(* Logix 5000 project; controller NWGG 1756-L72 rev 35.12; software revision 35.00; part 14 of 19 *)
(* tags used below, declared in another part *)
   ALM_Air_Gate_Failed_Open_Bin0 : ALARM_DIGITAL;
   ALM_Air_Gate_Failed_Open_Bin1 : ALARM_DIGITAL;
   ALM_Air_Gate_Failed_Open_Bin10 : ALARM_DIGITAL;
   ALM_Air_Gate_Failed_Open_Bin11 : ALARM_DIGITAL;
   ALM_Air_Gate_Failed_Open_Bin12 : ALARM_DIGITAL;
   ALM_Air_Gate_Failed_Open_Bin13 : ALARM_DIGITAL;
   ALM_Air_Gate_Failed_Open_Bin14 : ALARM_DIGITAL;
   ALM_Air_Gate_Failed_Open_Bin15 : ALARM_DIGITAL;
   ALM_Air_Gate_Failed_Open_Bin16 : ALARM_DIGITAL;
   ALM_Air_Gate_Failed_Open_Bin2 : ALARM_DIGITAL;
   ALM_Air_Gate_Failed_Open_Bin5 : ALARM_DIGITAL;
   ALM_Air_Gate_Failed_Open_Bin6 : ALARM_DIGITAL;
   ALM_Air_Gate_Failed_Open_Bin7 : ALARM_DIGITAL;
   ALM_Air_Gate_Failed_Open_Bin8 : ALARM_DIGITAL;
   ALM_Air_Gate_Failed_Open_Bin9 : ALARM_DIGITAL;
   ALM_OVRAMP_Belt10 : ALARM_DIGITAL;
   ALM_OVRAMP_Belt11 : ALARM_DIGITAL;
   ALM_OVRAMP_Belt2 : ALARM_DIGITAL;
   ALM_OVRAMP_Belt3 : ALARM_DIGITAL;
   ALM_OVRAMP_Belt5 : ALARM_DIGITAL;
   ALM_OVRAMP_Belt6 : ALARM_DIGITAL;
   ALM_OVRAMP_Belt7 : ALARM_DIGITAL;
   ALM_OVRAMP_Belt8 : ALARM_DIGITAL;
   ALM_OVRAMP_Belt9 : ALARM_DIGITAL;
   ALM_PLUG_Belt1 : ALARM_DIGITAL;
   ALM_PLUG_Belt10 : ALARM_DIGITAL;
   ALM_PLUG_Belt11 : ALARM_DIGITAL;
   ALM_PLUG_Belt2 : ALARM_DIGITAL;
   ALM_PLUG_Belt3 : ALARM_DIGITAL;
   ALM_PLUG_Belt5 : ALARM_DIGITAL;
   ALM_PLUG_Belt6 : ALARM_DIGITAL;
   ALM_PLUG_Belt7 : ALARM_DIGITAL;
   ALM_PLUG_Belt8 : ALARM_DIGITAL;
   ALM_PLUG_Belt9 : ALARM_DIGITAL;
   ALM_SLP10_Belt1 : ALARM_DIGITAL;
   ALM_SLP10_Belt10 : ALARM_DIGITAL;
   ALM_SLP10_Belt11 : ALARM_DIGITAL;
   ALM_SLP10_Belt2 : ALARM_DIGITAL;
   ALM_SLP10_Belt3 : ALARM_DIGITAL;
   ALM_SLP10_Belt5 : ALARM_DIGITAL;
   ALM_SLP10_Belt6 : ALARM_DIGITAL;
   ALM_SLP10_Belt7 : ALARM_DIGITAL;
   ALM_SLP10_Belt8 : ALARM_DIGITAL;
   ALM_SLP10_Belt9 : ALARM_DIGITAL;
   ALM_SLP20_Belt1 : ALARM_DIGITAL;
   ALM_SLP20_Belt10 : ALARM_DIGITAL;
   ALM_SLP20_Belt11 : ALARM_DIGITAL;
   ALM_SLP20_Belt2 : ALARM_DIGITAL;
   ALM_SLP20_Belt3 : ALARM_DIGITAL;
   ALM_SLP20_Belt5 : ALARM_DIGITAL;
   ALM_SLP20_Belt6 : ALARM_DIGITAL;
   ALM_SLP20_Belt7 : ALARM_DIGITAL;
   ALM_SLP20_Belt8 : ALARM_DIGITAL;
   ALM_SLP20_Belt9 : ALARM_DIGITAL;
   ALM_WONT_START_Belt1 : ALARM_DIGITAL;
   ALM_WONT_START_Belt10 : ALARM_DIGITAL;
   ALM_WONT_START_Belt11 : ALARM_DIGITAL;
   ALM_WONT_START_Belt2 : ALARM_DIGITAL;
   ALM_WONT_START_Belt3 : ALARM_DIGITAL;
   ALM_WONT_START_Belt5 : ALARM_DIGITAL;
   ALM_WONT_START_Belt6 : ALARM_DIGITAL;
   ALM_WONT_START_Belt7 : ALARM_DIGITAL;
   ALM_WONT_START_Belt8 : ALARM_DIGITAL;
   ALM_WONT_START_Belt9 : ALARM_DIGITAL;
   Always_Off : BOOL;
   Andco_Rate : DINT;
   b3 : ALARM_DIGITAL;
   Batch_Status : DINT;
   BC_9_Interlock : BOOL;
   Belt : udt_Motor[16];
   Bin_Clean_Pause : BOOL;
   Bin_Loadout_Control : Loadout_Bin_Control[29];
   Bin_Transfer_Pause : BOOL;
   Bin_Treat_Pause : BOOL;
   Clean_Batch_Status : DINT;
   Concrete_Leg : udt_Motor;
   Config_Bin_Name : STRING;
   Config_Cancel_Bin : BOOL;
   Config_Class : STRING;
   Config_Clean_Delay_Start : REAL;
   Config_Clean_Delay_Stop : REAL;
   Config_Item_Number : STRING;
   Config_Name : STRING;
   Config_Pounds_Per_Inch : REAL;
   Config_Save_Bin : BOOL;
   Config_Treat_Delay_Start : REAL;
   Config_Treat_Delay_Stop : REAL;
   ConfigureIndex : DINT;
   Empty_String : STRING;
   IDX : DINT;
   Interlock_Not_Used : BOOL;
   loa : ALARM_DIGITAL;
   Loadout_Bin : udt_Loadout_Bin[29];
   Loadout_K_Valve : udt_Loadout_K_Valve[2];
   Man_Start_Stop_Allowed : BOOL;
   Manual_Mode : BOOL;
   Move_Bin_Config : BOOL;
   NA : BOOL;
   TMR_Max_Clean_Delay : TIMER;
   TMR_Max_Treat_Delay : TIMER;
   Transfer_Batch_Status : DINT;
   Treat_Batch_Status : DINT;
   Treater_Loadout : udt_Treater_Loadout;
   _700_AIR_GA : ALIAS FOR I8.3;
   _700G_CLOSE : ALIAS FOR O12.9;
   _700G_OPEN : ALIAS FOR O12.8;
   _701_AIR_GA : ALIAS FOR I8.5;
   Always_On : BOOL;
   Bin_Config : BOOL;
   CP_Remote_Air_Gate_On : DINT;
   CP_Remote_Air_Gate_Open_In : DINT;
   CP_Remote_Andoc_Out : udt_Andco_Remote_Out[32];
   CP_Remote_Belt_In : udt_Motor_Remote_In[10];
   CP_Remote_Belt_Start : DINT;
   I1_000_Bit00 : ALIAS FOR I1.0;
   I4_000_Bit11 : ALIAS FOR I4.11;
   I8_000_Bit08 : ALIAS FOR I8.8;
   I8_000_Bit09 : ALIAS FOR I8.9;
   I8_000_Bit10 : ALIAS FOR I8.10;
   I8_000_Bit11 : ALIAS FOR I8.11;
   O12_000_Bit10 : ALIAS FOR O12.10;
   O12_000_Bit11 : ALIAS FOR O12.11;
   O12_000_Bit12 : ALIAS FOR O12.12;
   O12_000_Bit13 : ALIAS FOR O12.13;
   O9_000_Bit00 : ALIAS FOR O9.0;
   O9_000_Bit01 : ALIAS FOR O9.1;
   O9_000_Bit02 : ALIAS FOR O9.2;
   RemoteAndcoAnalogIn : DINT[40];
(* SeedLoadoutMain, continued *)

ROUTINE Amp_Gages   (* function block diagram *)
   SHEET 1
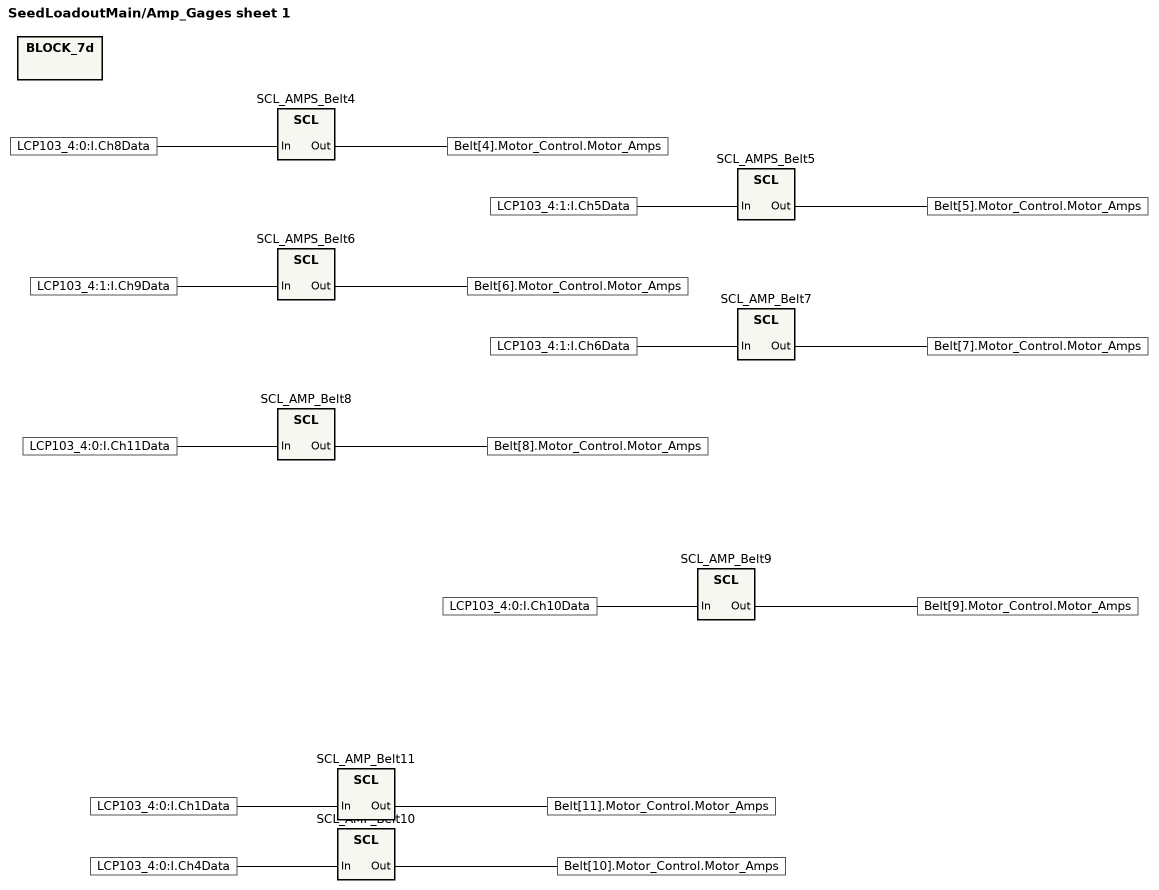
   BLOCK_7d_1 : BLOCK_7d();
   SCL_AMPS_Belt4 : SCL(In := LCP103_4:0:I.Ch8Data);
   SCL_AMPS_Belt6 : SCL(In := LCP103_4:1:I.Ch9Data);
   SCL_AMP_Belt8 : SCL(In := LCP103_4:0:I.Ch11Data);
   SCL_AMP_Belt11 : SCL(In := LCP103_4:0:I.Ch1Data);
   SCL_AMP_Belt10 : SCL(In := LCP103_4:0:I.Ch4Data);
   Belt[4].Motor_Control.Motor_Amps := SCL_AMPS_Belt4.Out;
   Belt[6].Motor_Control.Motor_Amps := SCL_AMPS_Belt6.Out;
   Belt[8].Motor_Control.Motor_Amps := SCL_AMP_Belt8.Out;
   Belt[11].Motor_Control.Motor_Amps := SCL_AMP_Belt11.Out;
   Belt[10].Motor_Control.Motor_Amps := SCL_AMP_Belt10.Out;
   SCL_AMP_Belt9 : SCL(In := LCP103_4:0:I.Ch10Data);
   SCL_AMPS_Belt5 : SCL(In := LCP103_4:1:I.Ch5Data);
   SCL_AMP_Belt7 : SCL(In := LCP103_4:1:I.Ch6Data);
   Belt[9].Motor_Control.Motor_Amps := SCL_AMP_Belt9.Out;
   Belt[5].Motor_Control.Motor_Amps := SCL_AMPS_Belt5.Out;
   Belt[7].Motor_Control.Motor_Amps := SCL_AMP_Belt7.Out;
END_ROUTINE

ROUTINE Andco_Rate   (* ladder *)
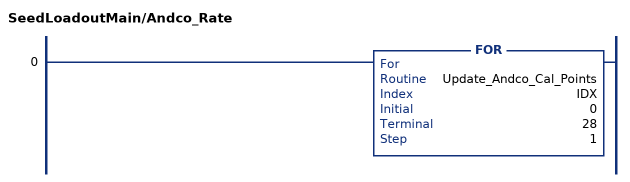
   0: FOR(Update_Andco_Cal_Points,IDX,0,28,1);
END_ROUTINE

ROUTINE Batch_Status   (* ladder *)
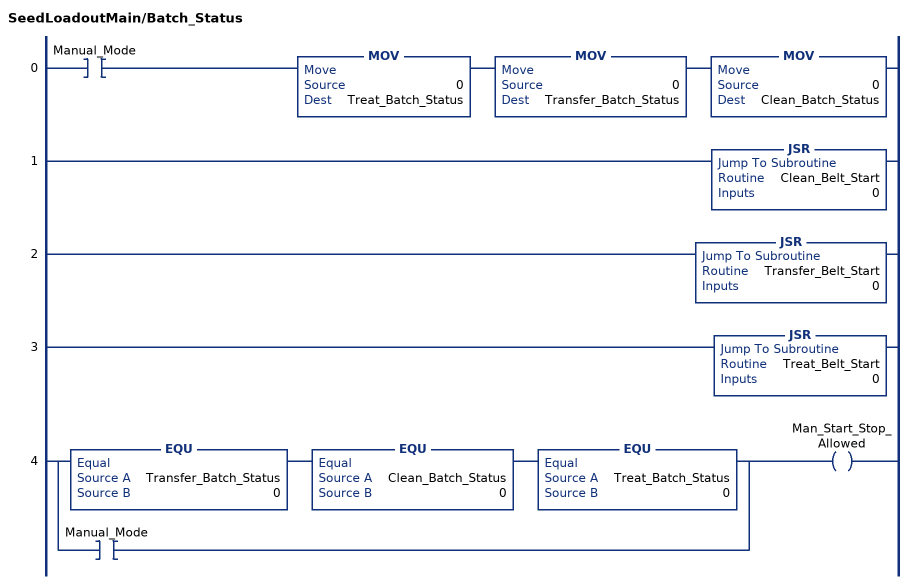
   0: XIC(Manual_Mode)MOV(0,Treat_Batch_Status)MOV(0,Transfer_Batch_Status)MOV(0,Clean_Batch_Status);
   1: JSR(Clean_Belt_Start,0);
   2: JSR(Transfer_Belt_Start,0);
   3: JSR(Treat_Belt_Start,0);
   4: [EQU(Transfer_Batch_Status,0) EQU(Clean_Batch_Status,0) EQU(Treat_Batch_Status,0) ,XIC(Manual_Mode) ]OTE(Man_Start_Stop_Allowed);
END_ROUTINE

ROUTINE Belts   (* ladder *)
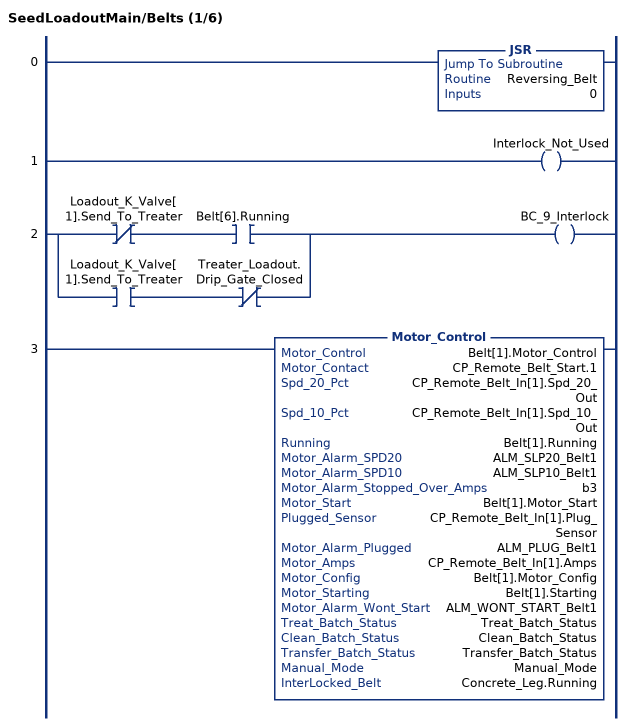
   0: JSR(Reversing_Belt,0);
   1: OTE(Interlock_Not_Used);
   2: [XIO(Loadout_K_Valve[1].Send_To_Treater) XIC(Belt[6].Running) ,XIC(Loadout_K_Valve[1].Send_To_Treater) XIO(Treater_Loadout.Drip_Gate_Closed) ]OTE(BC_9_Interlock);
   3: Motor_Control(Belt[1].Motor_Control,CP_Remote_Belt_Start.1,CP_Remote_Belt_In[1].Spd_20_Out,CP_Remote_Belt_In[1].Spd_10_Out,Belt[1].Running,ALM_SLP20_Belt1,ALM_SLP10_Belt1,b3,Belt[1].Motor_Start,CP_Remote_Belt_In[1].Plug_Sensor,ALM_PLUG_Belt1,CP_Remote_Belt_In[1].Amps,Belt[1].Motor_Config,Belt[1].Starting,ALM_WONT_START_Belt1,Treat_Batch_Status,Clean_Batch_Status,Transfer_Batch_Status,Manual_Mode,Concrete_Leg.Running);
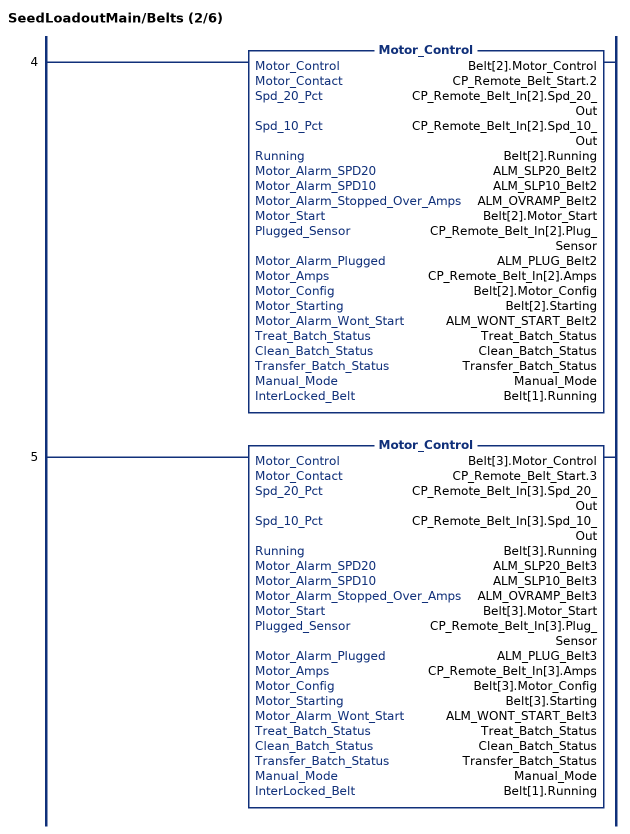
   4: Motor_Control(Belt[2].Motor_Control,CP_Remote_Belt_Start.2,CP_Remote_Belt_In[2].Spd_20_Out,CP_Remote_Belt_In[2].Spd_10_Out,Belt[2].Running,ALM_SLP20_Belt2,ALM_SLP10_Belt2,ALM_OVRAMP_Belt2,Belt[2].Motor_Start,CP_Remote_Belt_In[2].Plug_Sensor,ALM_PLUG_Belt2,CP_Remote_Belt_In[2].Amps,Belt[2].Motor_Config,Belt[2].Starting,ALM_WONT_START_Belt2,Treat_Batch_Status,Clean_Batch_Status,Transfer_Batch_Status,Manual_Mode,Belt[1].Running);
   5: Motor_Control(Belt[3].Motor_Control,CP_Remote_Belt_Start.3,CP_Remote_Belt_In[3].Spd_20_Out,CP_Remote_Belt_In[3].Spd_10_Out,Belt[3].Running,ALM_SLP20_Belt3,ALM_SLP10_Belt3,ALM_OVRAMP_Belt3,Belt[3].Motor_Start,CP_Remote_Belt_In[3].Plug_Sensor,ALM_PLUG_Belt3,CP_Remote_Belt_In[3].Amps,Belt[3].Motor_Config,Belt[3].Starting,ALM_WONT_START_Belt3,Treat_Batch_Status,Clean_Batch_Status,Transfer_Batch_Status,Manual_Mode,Belt[1].Running);
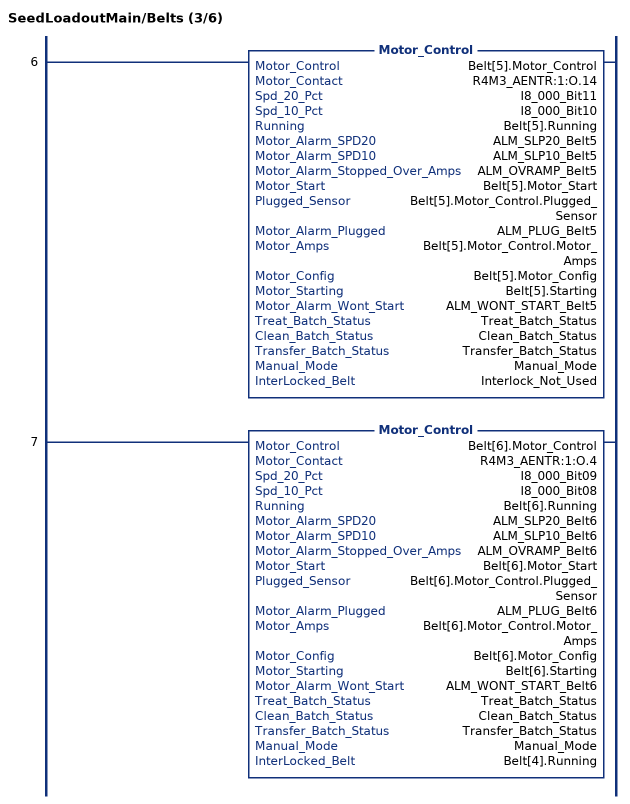
   6: Motor_Control(Belt[5].Motor_Control,R4M3_AENTR:1:O.14,I8_000_Bit11,I8_000_Bit10,Belt[5].Running,ALM_SLP20_Belt5,ALM_SLP10_Belt5,ALM_OVRAMP_Belt5,Belt[5].Motor_Start,Belt[5].Motor_Control.Plugged_Sensor,ALM_PLUG_Belt5,Belt[5].Motor_Control.Motor_Amps,Belt[5].Motor_Config,Belt[5].Starting,ALM_WONT_START_Belt5,Treat_Batch_Status,Clean_Batch_Status,Transfer_Batch_Status,Manual_Mode,Interlock_Not_Used);
   7: Motor_Control(Belt[6].Motor_Control,R4M3_AENTR:1:O.4,I8_000_Bit09,I8_000_Bit08,Belt[6].Running,ALM_SLP20_Belt6,ALM_SLP10_Belt6,ALM_OVRAMP_Belt6,Belt[6].Motor_Start,Belt[6].Motor_Control.Plugged_Sensor,ALM_PLUG_Belt6,Belt[6].Motor_Control.Motor_Amps,Belt[6].Motor_Config,Belt[6].Starting,ALM_WONT_START_Belt6,Treat_Batch_Status,Clean_Batch_Status,Transfer_Batch_Status,Manual_Mode,Belt[4].Running);
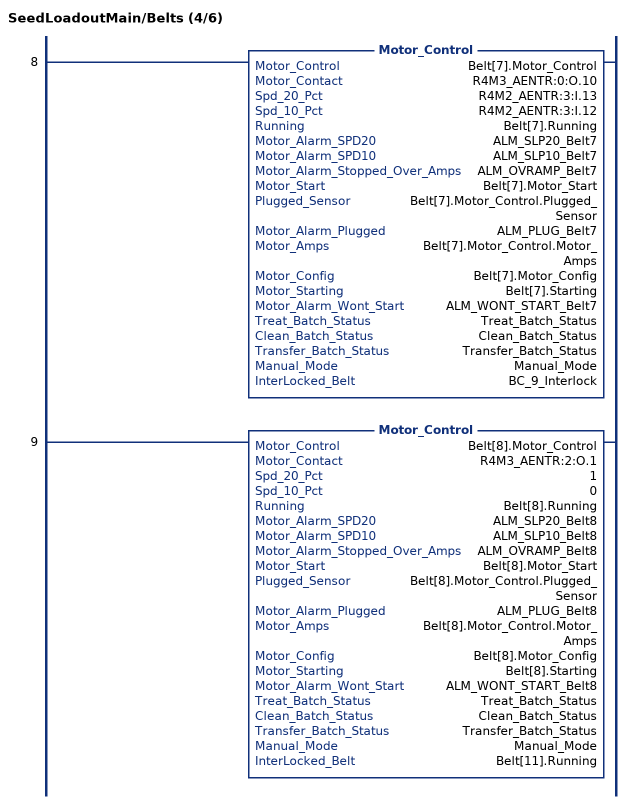
   8: Motor_Control(Belt[7].Motor_Control,R4M3_AENTR:0:O.10,R4M2_AENTR:3:I.13,R4M2_AENTR:3:I.12,Belt[7].Running,ALM_SLP20_Belt7,ALM_SLP10_Belt7,ALM_OVRAMP_Belt7,Belt[7].Motor_Start,Belt[7].Motor_Control.Plugged_Sensor,ALM_PLUG_Belt7,Belt[7].Motor_Control.Motor_Amps,Belt[7].Motor_Config,Belt[7].Starting,ALM_WONT_START_Belt7,Treat_Batch_Status,Clean_Batch_Status,Transfer_Batch_Status,Manual_Mode,BC_9_Interlock);
   9: Motor_Control(Belt[8].Motor_Control,R4M3_AENTR:2:O.1,1,0,Belt[8].Running,ALM_SLP20_Belt8,ALM_SLP10_Belt8,ALM_OVRAMP_Belt8,Belt[8].Motor_Start,Belt[8].Motor_Control.Plugged_Sensor,ALM_PLUG_Belt8,Belt[8].Motor_Control.Motor_Amps,Belt[8].Motor_Config,Belt[8].Starting,ALM_WONT_START_Belt8,Treat_Batch_Status,Clean_Batch_Status,Transfer_Batch_Status,Manual_Mode,Belt[11].Running);
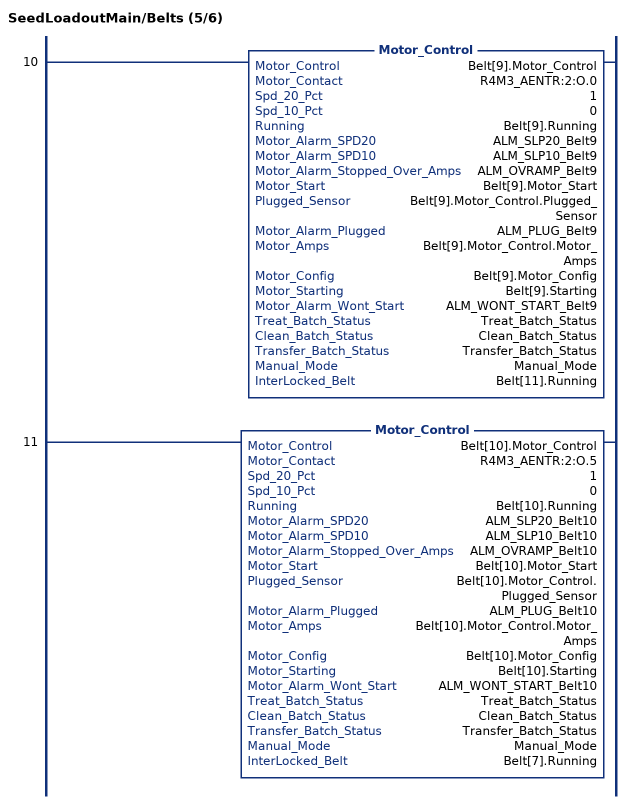
   10: Motor_Control(Belt[9].Motor_Control,R4M3_AENTR:2:O.0,1,0,Belt[9].Running,ALM_SLP20_Belt9,ALM_SLP10_Belt9,ALM_OVRAMP_Belt9,Belt[9].Motor_Start,Belt[9].Motor_Control.Plugged_Sensor,ALM_PLUG_Belt9,Belt[9].Motor_Control.Motor_Amps,Belt[9].Motor_Config,Belt[9].Starting,ALM_WONT_START_Belt9,Treat_Batch_Status,Clean_Batch_Status,Transfer_Batch_Status,Manual_Mode,Belt[11].Running);
   11: Motor_Control(Belt[10].Motor_Control,R4M3_AENTR:2:O.5,1,0,Belt[10].Running,ALM_SLP20_Belt10,ALM_SLP10_Belt10,ALM_OVRAMP_Belt10,Belt[10].Motor_Start,Belt[10].Motor_Control.Plugged_Sensor,ALM_PLUG_Belt10,Belt[10].Motor_Control.Motor_Amps,Belt[10].Motor_Config,Belt[10].Starting,ALM_WONT_START_Belt10,Treat_Batch_Status,Clean_Batch_Status,Transfer_Batch_Status,Manual_Mode,Belt[7].Running);
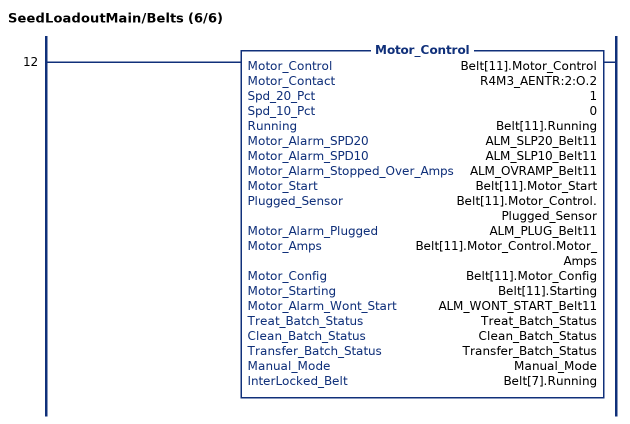
   12: Motor_Control(Belt[11].Motor_Control,R4M3_AENTR:2:O.2,1,0,Belt[11].Running,ALM_SLP20_Belt11,ALM_SLP10_Belt11,ALM_OVRAMP_Belt11,Belt[11].Motor_Start,Belt[11].Motor_Control.Plugged_Sensor,ALM_PLUG_Belt11,Belt[11].Motor_Control.Motor_Amps,Belt[11].Motor_Config,Belt[11].Starting,ALM_WONT_START_Belt11,Treat_Batch_Status,Clean_Batch_Status,Transfer_Batch_Status,Manual_Mode,Belt[7].Running);
END_ROUTINE

ROUTINE BinConfigure   (* ladder *)
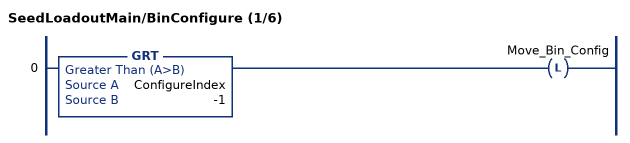
   0: GRT(ConfigureIndex,-1)OTL(Move_Bin_Config);
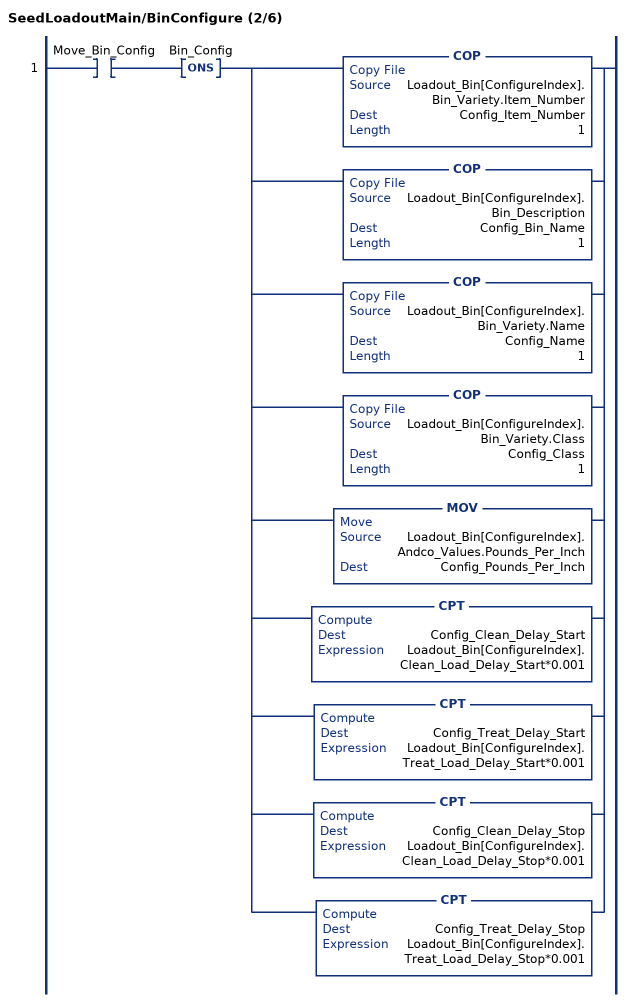
   1: XIC(Move_Bin_Config)ONS(Bin_Config)[COP(Loadout_Bin[ConfigureIndex].Bin_Variety.Item_Number,Config_Item_Number,1) ,COP(Loadout_Bin[ConfigureIndex].Bin_Description,Config_Bin_Name,1) ,COP(Loadout_Bin[ConfigureIndex].Bin_Variety.Name,Config_Name,1) ,COP(Loadout_Bin[ConfigureIndex].Bin_Variety.Class,Config_Class,1) ,MOV(Loadout_Bin[ConfigureIndex].Andco_Values.Pounds_Per_Inch,Config_Pounds_Per_Inch) ,CPT(Config_Clean_Delay_Start,Loadout_Bin[ConfigureIndex].Clean_Load_Delay_Start*0.001) ,CPT(Config_Treat_Delay_Start,Loadout_Bin[ConfigureIndex].Treat_Load_Delay_Start*0.001) ,CPT(Config_Clean_Delay_Stop,Loadout_Bin[ConfigureIndex].Clean_Load_Delay_Stop*0.001) ,CPT(Config_Treat_Delay_Stop,Loadout_Bin[ConfigureIndex].Treat_Load_Delay_Stop*0.001) ];
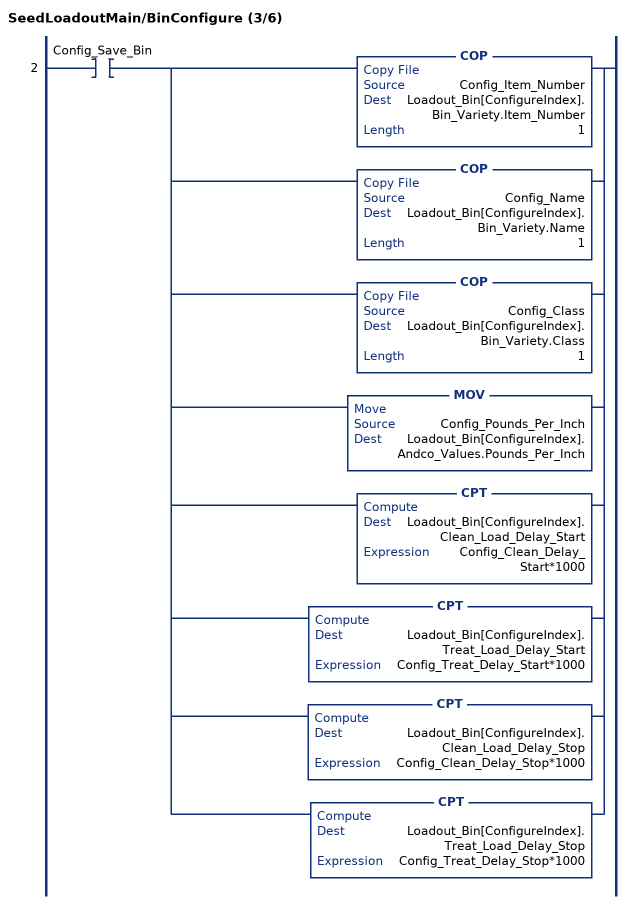
   2: XIC(Config_Save_Bin)[COP(Config_Item_Number,Loadout_Bin[ConfigureIndex].Bin_Variety.Item_Number,1) ,COP(Config_Name,Loadout_Bin[ConfigureIndex].Bin_Variety.Name,1) ,COP(Config_Class,Loadout_Bin[ConfigureIndex].Bin_Variety.Class,1) ,MOV(Config_Pounds_Per_Inch,Loadout_Bin[ConfigureIndex].Andco_Values.Pounds_Per_Inch) ,CPT(Loadout_Bin[ConfigureIndex].Clean_Load_Delay_Start,Config_Clean_Delay_Start*1000) ,CPT(Loadout_Bin[ConfigureIndex].Treat_Load_Delay_Start,Config_Treat_Delay_Start*1000) ,CPT(Loadout_Bin[ConfigureIndex].Clean_Load_Delay_Stop,Config_Clean_Delay_Stop*1000) ,CPT(Loadout_Bin[ConfigureIndex].Treat_Load_Delay_Stop,Config_Treat_Delay_Stop*1000) ];
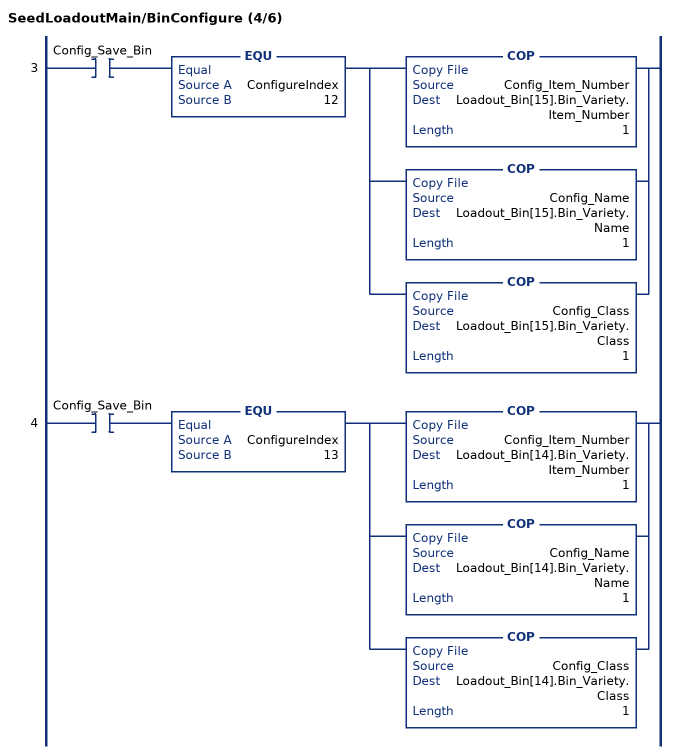
   3: XIC(Config_Save_Bin)EQU(ConfigureIndex,12)[COP(Config_Item_Number,Loadout_Bin[15].Bin_Variety.Item_Number,1) ,[COP(Config_Name,Loadout_Bin[15].Bin_Variety.Name,1) ,COP(Config_Class,Loadout_Bin[15].Bin_Variety.Class,1) ] ];
   4: XIC(Config_Save_Bin)EQU(ConfigureIndex,13)[COP(Config_Item_Number,Loadout_Bin[14].Bin_Variety.Item_Number,1) ,[COP(Config_Name,Loadout_Bin[14].Bin_Variety.Name,1) ,COP(Config_Class,Loadout_Bin[14].Bin_Variety.Class,1) ] ];
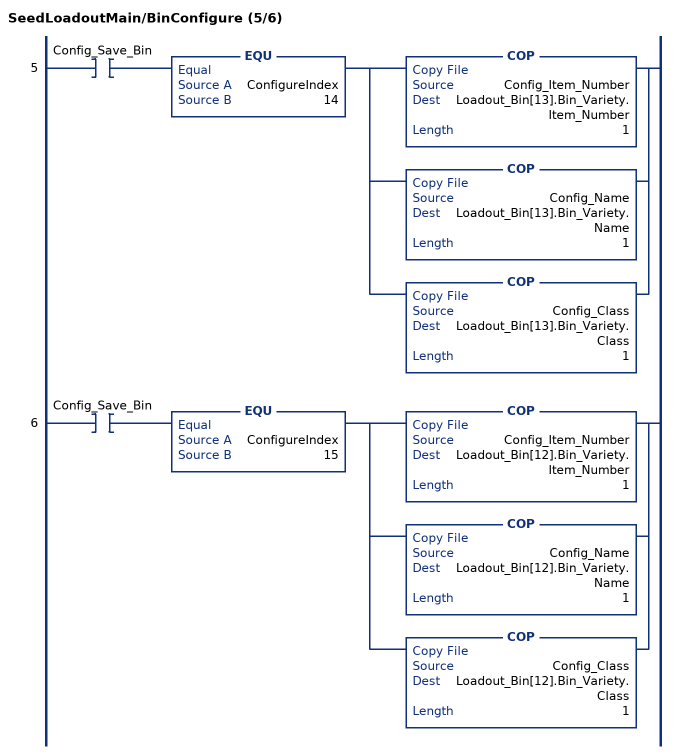
   5: XIC(Config_Save_Bin)EQU(ConfigureIndex,14)[COP(Config_Item_Number,Loadout_Bin[13].Bin_Variety.Item_Number,1) ,[COP(Config_Name,Loadout_Bin[13].Bin_Variety.Name,1) ,COP(Config_Class,Loadout_Bin[13].Bin_Variety.Class,1) ] ];
   6: XIC(Config_Save_Bin)EQU(ConfigureIndex,15)[COP(Config_Item_Number,Loadout_Bin[12].Bin_Variety.Item_Number,1) ,[COP(Config_Name,Loadout_Bin[12].Bin_Variety.Name,1) ,COP(Config_Class,Loadout_Bin[12].Bin_Variety.Class,1) ] ];
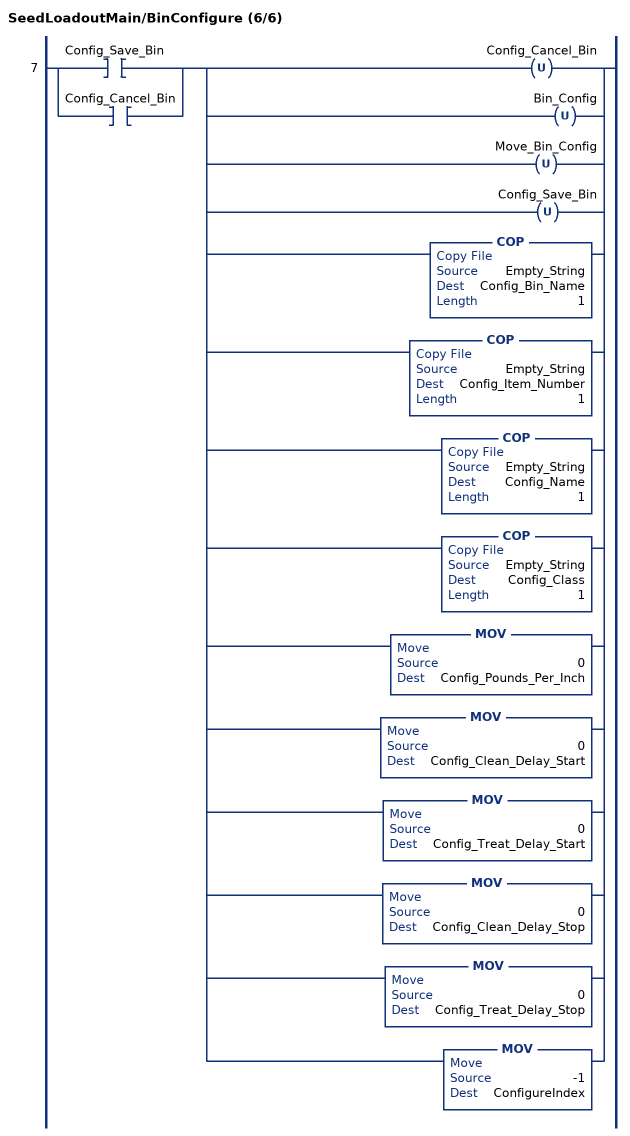
   7: [XIC(Config_Save_Bin) ,XIC(Config_Cancel_Bin) ][OTU(Config_Cancel_Bin) ,OTU(Bin_Config) ,OTU(Move_Bin_Config) ,OTU(Config_Save_Bin) ,COP(Empty_String,Config_Bin_Name,1) ,COP(Empty_String,Config_Item_Number,1) ,COP(Empty_String,Config_Name,1) ,COP(Empty_String,Config_Class,1) ,MOV(0,Config_Pounds_Per_Inch) ,MOV(0,Config_Clean_Delay_Start) ,MOV(0,Config_Treat_Delay_Start) ,MOV(0,Config_Clean_Delay_Stop) ,MOV(0,Config_Treat_Delay_Stop) ,MOV(-1,ConfigureIndex) ];
END_ROUTINE

ROUTINE Bins   (* ladder *)
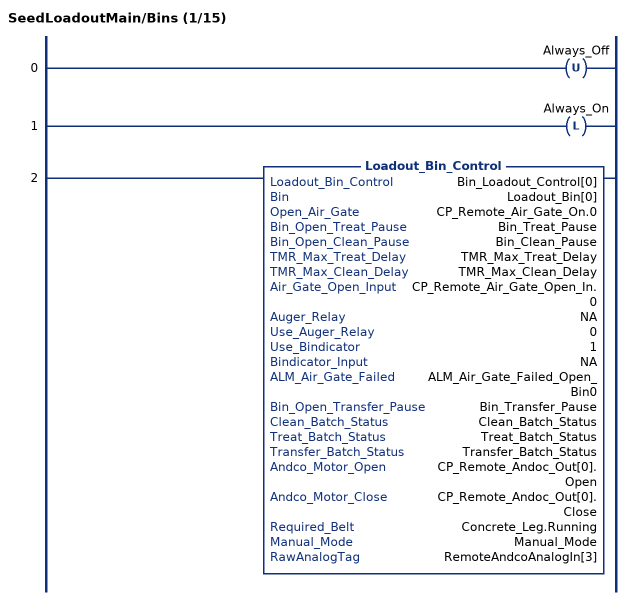
   0: OTU(Always_Off);
   1: OTL(Always_On);
   2: Loadout_Bin_Control(Bin_Loadout_Control[0],Loadout_Bin[0],CP_Remote_Air_Gate_On.0,Bin_Treat_Pause,Bin_Clean_Pause,TMR_Max_Treat_Delay,TMR_Max_Clean_Delay,CP_Remote_Air_Gate_Open_In.0,NA,0,1,NA,ALM_Air_Gate_Failed_Open_Bin0,Bin_Transfer_Pause,Clean_Batch_Status,Treat_Batch_Status,Transfer_Batch_Status,CP_Remote_Andoc_Out[0].Open,CP_Remote_Andoc_Out[0].Close,Concrete_Leg.Running,Manual_Mode,RemoteAndcoAnalogIn[3]);
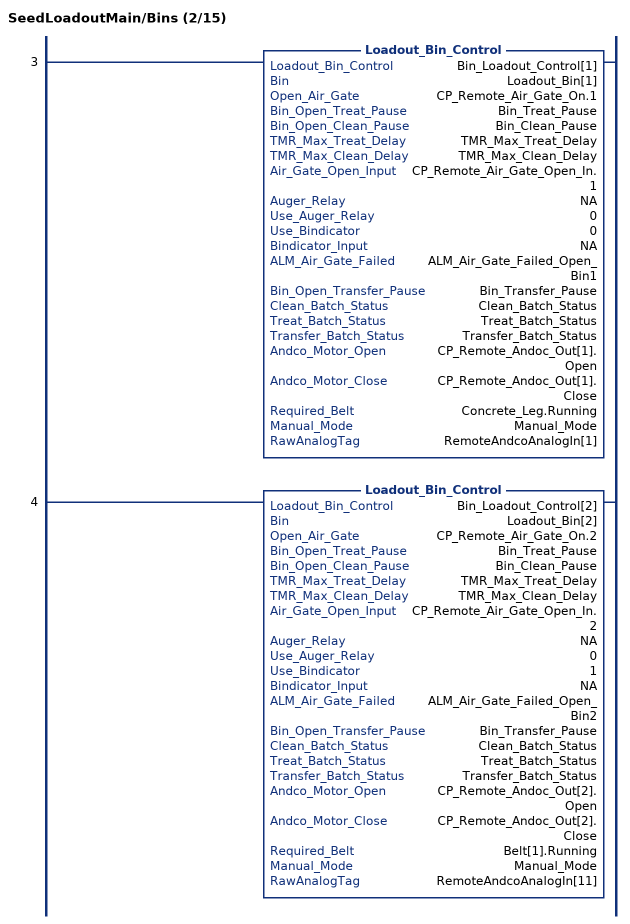
   3: Loadout_Bin_Control(Bin_Loadout_Control[1],Loadout_Bin[1],CP_Remote_Air_Gate_On.1,Bin_Treat_Pause,Bin_Clean_Pause,TMR_Max_Treat_Delay,TMR_Max_Clean_Delay,CP_Remote_Air_Gate_Open_In.1,NA,0,0,NA,ALM_Air_Gate_Failed_Open_Bin1,Bin_Transfer_Pause,Clean_Batch_Status,Treat_Batch_Status,Transfer_Batch_Status,CP_Remote_Andoc_Out[1].Open,CP_Remote_Andoc_Out[1].Close,Concrete_Leg.Running,Manual_Mode,RemoteAndcoAnalogIn[1]);
   4: Loadout_Bin_Control(Bin_Loadout_Control[2],Loadout_Bin[2],CP_Remote_Air_Gate_On.2,Bin_Treat_Pause,Bin_Clean_Pause,TMR_Max_Treat_Delay,TMR_Max_Clean_Delay,CP_Remote_Air_Gate_Open_In.2,NA,0,1,NA,ALM_Air_Gate_Failed_Open_Bin2,Bin_Transfer_Pause,Clean_Batch_Status,Treat_Batch_Status,Transfer_Batch_Status,CP_Remote_Andoc_Out[2].Open,CP_Remote_Andoc_Out[2].Close,Belt[1].Running,Manual_Mode,RemoteAndcoAnalogIn[11]);
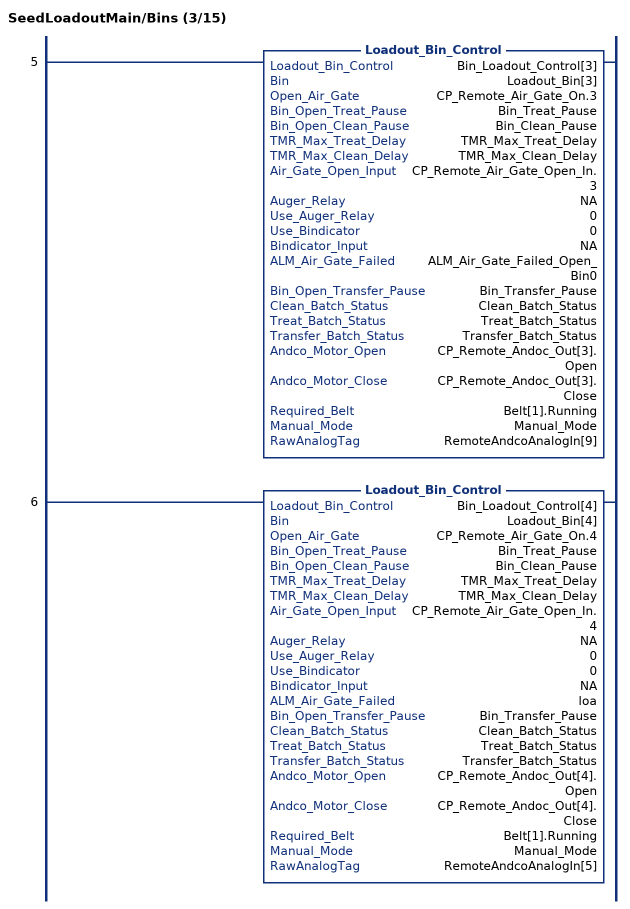
   5: Loadout_Bin_Control(Bin_Loadout_Control[3],Loadout_Bin[3],CP_Remote_Air_Gate_On.3,Bin_Treat_Pause,Bin_Clean_Pause,TMR_Max_Treat_Delay,TMR_Max_Clean_Delay,CP_Remote_Air_Gate_Open_In.3,NA,0,0,NA,ALM_Air_Gate_Failed_Open_Bin0,Bin_Transfer_Pause,Clean_Batch_Status,Treat_Batch_Status,Transfer_Batch_Status,CP_Remote_Andoc_Out[3].Open,CP_Remote_Andoc_Out[3].Close,Belt[1].Running,Manual_Mode,RemoteAndcoAnalogIn[9]);
   6: Loadout_Bin_Control(Bin_Loadout_Control[4],Loadout_Bin[4],CP_Remote_Air_Gate_On.4,Bin_Treat_Pause,Bin_Clean_Pause,TMR_Max_Treat_Delay,TMR_Max_Clean_Delay,CP_Remote_Air_Gate_Open_In.4,NA,0,0,NA,loa,Bin_Transfer_Pause,Clean_Batch_Status,Treat_Batch_Status,Transfer_Batch_Status,CP_Remote_Andoc_Out[4].Open,CP_Remote_Andoc_Out[4].Close,Belt[1].Running,Manual_Mode,RemoteAndcoAnalogIn[5]);
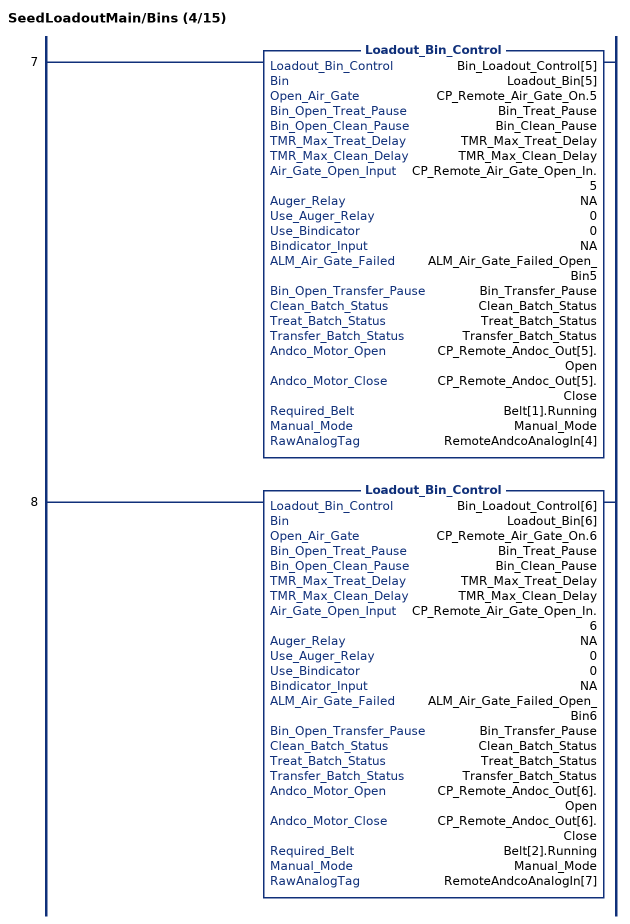
   7: Loadout_Bin_Control(Bin_Loadout_Control[5],Loadout_Bin[5],CP_Remote_Air_Gate_On.5,Bin_Treat_Pause,Bin_Clean_Pause,TMR_Max_Treat_Delay,TMR_Max_Clean_Delay,CP_Remote_Air_Gate_Open_In.5,NA,0,0,NA,ALM_Air_Gate_Failed_Open_Bin5,Bin_Transfer_Pause,Clean_Batch_Status,Treat_Batch_Status,Transfer_Batch_Status,CP_Remote_Andoc_Out[5].Open,CP_Remote_Andoc_Out[5].Close,Belt[1].Running,Manual_Mode,RemoteAndcoAnalogIn[4]);
   8: Loadout_Bin_Control(Bin_Loadout_Control[6],Loadout_Bin[6],CP_Remote_Air_Gate_On.6,Bin_Treat_Pause,Bin_Clean_Pause,TMR_Max_Treat_Delay,TMR_Max_Clean_Delay,CP_Remote_Air_Gate_Open_In.6,NA,0,0,NA,ALM_Air_Gate_Failed_Open_Bin6,Bin_Transfer_Pause,Clean_Batch_Status,Treat_Batch_Status,Transfer_Batch_Status,CP_Remote_Andoc_Out[6].Open,CP_Remote_Andoc_Out[6].Close,Belt[2].Running,Manual_Mode,RemoteAndcoAnalogIn[7]);
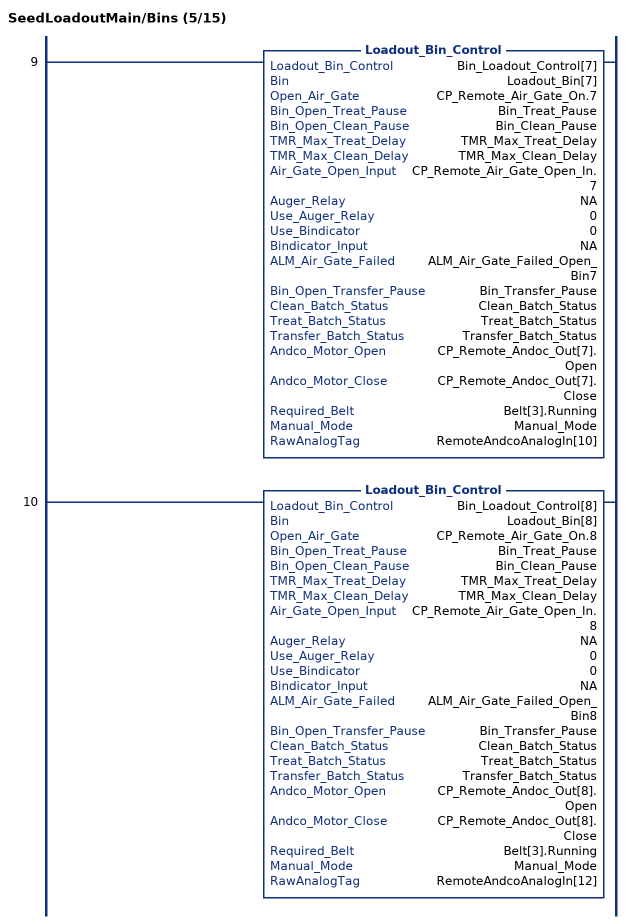
   9: Loadout_Bin_Control(Bin_Loadout_Control[7],Loadout_Bin[7],CP_Remote_Air_Gate_On.7,Bin_Treat_Pause,Bin_Clean_Pause,TMR_Max_Treat_Delay,TMR_Max_Clean_Delay,CP_Remote_Air_Gate_Open_In.7,NA,0,0,NA,ALM_Air_Gate_Failed_Open_Bin7,Bin_Transfer_Pause,Clean_Batch_Status,Treat_Batch_Status,Transfer_Batch_Status,CP_Remote_Andoc_Out[7].Open,CP_Remote_Andoc_Out[7].Close,Belt[3].Running,Manual_Mode,RemoteAndcoAnalogIn[10]);
   10: Loadout_Bin_Control(Bin_Loadout_Control[8],Loadout_Bin[8],CP_Remote_Air_Gate_On.8,Bin_Treat_Pause,Bin_Clean_Pause,TMR_Max_Treat_Delay,TMR_Max_Clean_Delay,CP_Remote_Air_Gate_Open_In.8,NA,0,0,NA,ALM_Air_Gate_Failed_Open_Bin8,Bin_Transfer_Pause,Clean_Batch_Status,Treat_Batch_Status,Transfer_Batch_Status,CP_Remote_Andoc_Out[8].Open,CP_Remote_Andoc_Out[8].Close,Belt[3].Running,Manual_Mode,RemoteAndcoAnalogIn[12]);
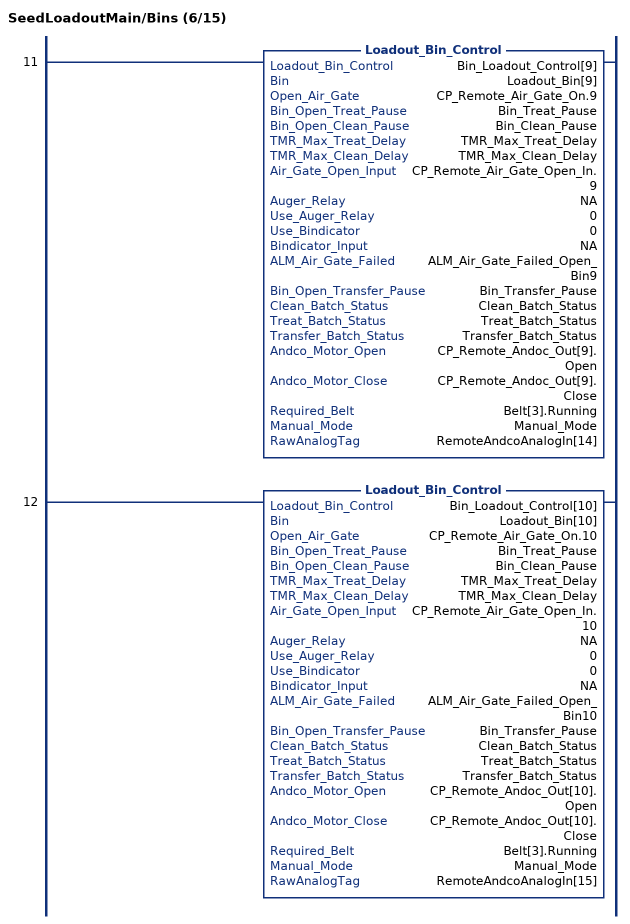
   11: Loadout_Bin_Control(Bin_Loadout_Control[9],Loadout_Bin[9],CP_Remote_Air_Gate_On.9,Bin_Treat_Pause,Bin_Clean_Pause,TMR_Max_Treat_Delay,TMR_Max_Clean_Delay,CP_Remote_Air_Gate_Open_In.9,NA,0,0,NA,ALM_Air_Gate_Failed_Open_Bin9,Bin_Transfer_Pause,Clean_Batch_Status,Treat_Batch_Status,Transfer_Batch_Status,CP_Remote_Andoc_Out[9].Open,CP_Remote_Andoc_Out[9].Close,Belt[3].Running,Manual_Mode,RemoteAndcoAnalogIn[14]);
   12: Loadout_Bin_Control(Bin_Loadout_Control[10],Loadout_Bin[10],CP_Remote_Air_Gate_On.10,Bin_Treat_Pause,Bin_Clean_Pause,TMR_Max_Treat_Delay,TMR_Max_Clean_Delay,CP_Remote_Air_Gate_Open_In.10,NA,0,0,NA,ALM_Air_Gate_Failed_Open_Bin10,Bin_Transfer_Pause,Clean_Batch_Status,Treat_Batch_Status,Transfer_Batch_Status,CP_Remote_Andoc_Out[10].Open,CP_Remote_Andoc_Out[10].Close,Belt[3].Running,Manual_Mode,RemoteAndcoAnalogIn[15]);
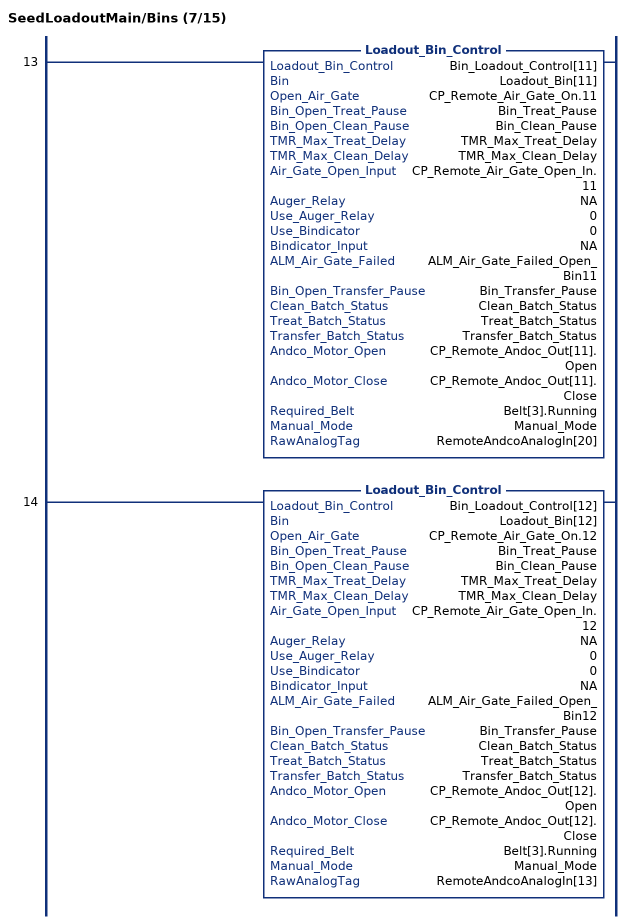
   13: Loadout_Bin_Control(Bin_Loadout_Control[11],Loadout_Bin[11],CP_Remote_Air_Gate_On.11,Bin_Treat_Pause,Bin_Clean_Pause,TMR_Max_Treat_Delay,TMR_Max_Clean_Delay,CP_Remote_Air_Gate_Open_In.11,NA,0,0,NA,ALM_Air_Gate_Failed_Open_Bin11,Bin_Transfer_Pause,Clean_Batch_Status,Treat_Batch_Status,Transfer_Batch_Status,CP_Remote_Andoc_Out[11].Open,CP_Remote_Andoc_Out[11].Close,Belt[3].Running,Manual_Mode,RemoteAndcoAnalogIn[20]);
   14: Loadout_Bin_Control(Bin_Loadout_Control[12],Loadout_Bin[12],CP_Remote_Air_Gate_On.12,Bin_Treat_Pause,Bin_Clean_Pause,TMR_Max_Treat_Delay,TMR_Max_Clean_Delay,CP_Remote_Air_Gate_Open_In.12,NA,0,0,NA,ALM_Air_Gate_Failed_Open_Bin12,Bin_Transfer_Pause,Clean_Batch_Status,Treat_Batch_Status,Transfer_Batch_Status,CP_Remote_Andoc_Out[12].Open,CP_Remote_Andoc_Out[12].Close,Belt[3].Running,Manual_Mode,RemoteAndcoAnalogIn[13]);
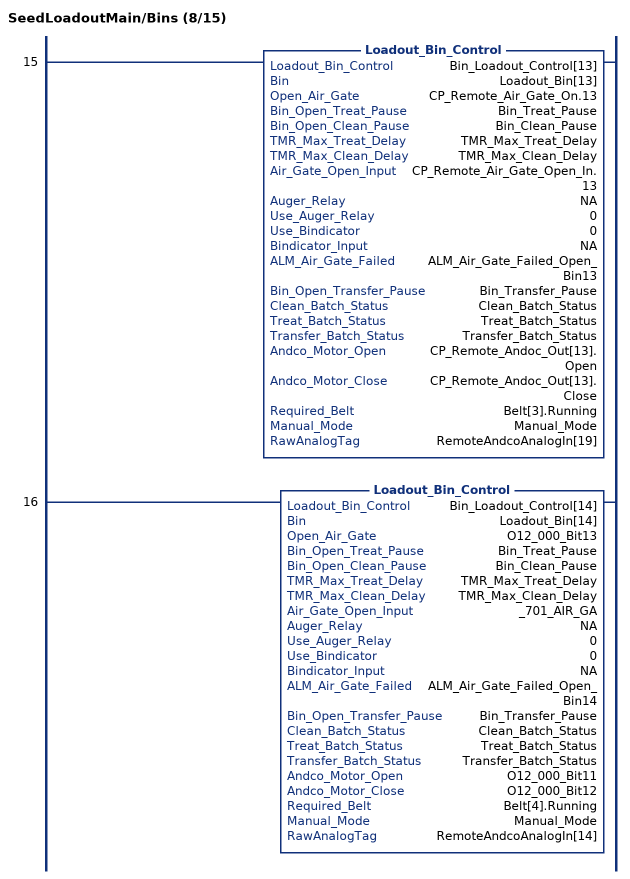
   15: Loadout_Bin_Control(Bin_Loadout_Control[13],Loadout_Bin[13],CP_Remote_Air_Gate_On.13,Bin_Treat_Pause,Bin_Clean_Pause,TMR_Max_Treat_Delay,TMR_Max_Clean_Delay,CP_Remote_Air_Gate_Open_In.13,NA,0,0,NA,ALM_Air_Gate_Failed_Open_Bin13,Bin_Transfer_Pause,Clean_Batch_Status,Treat_Batch_Status,Transfer_Batch_Status,CP_Remote_Andoc_Out[13].Open,CP_Remote_Andoc_Out[13].Close,Belt[3].Running,Manual_Mode,RemoteAndcoAnalogIn[19]);
   16: Loadout_Bin_Control(Bin_Loadout_Control[14],Loadout_Bin[14],O12_000_Bit13,Bin_Treat_Pause,Bin_Clean_Pause,TMR_Max_Treat_Delay,TMR_Max_Clean_Delay,_701_AIR_GA,NA,0,0,NA,ALM_Air_Gate_Failed_Open_Bin14,Bin_Transfer_Pause,Clean_Batch_Status,Treat_Batch_Status,Transfer_Batch_Status,O12_000_Bit11,O12_000_Bit12,Belt[4].Running,Manual_Mode,RemoteAndcoAnalogIn[14]);
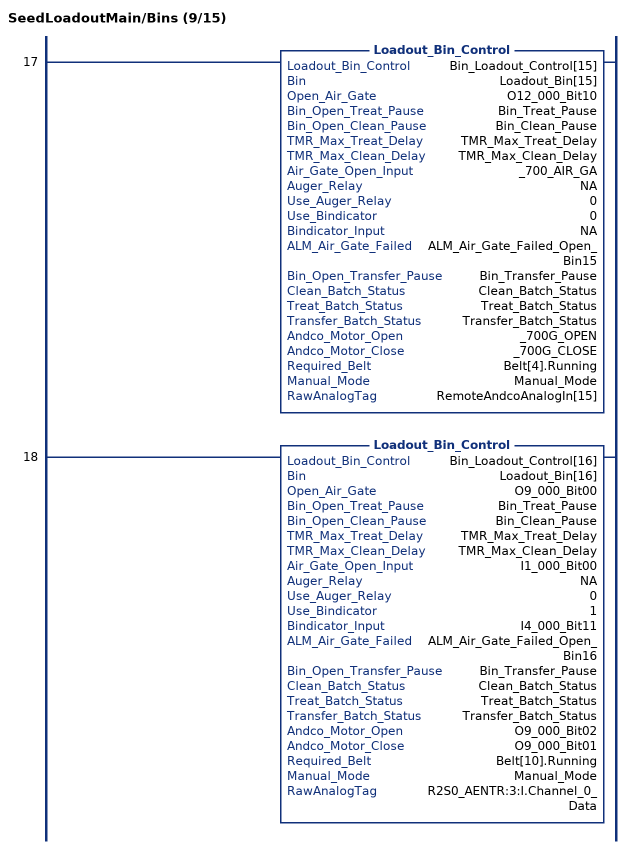
   17: Loadout_Bin_Control(Bin_Loadout_Control[15],Loadout_Bin[15],O12_000_Bit10,Bin_Treat_Pause,Bin_Clean_Pause,TMR_Max_Treat_Delay,TMR_Max_Clean_Delay,_700_AIR_GA,NA,0,0,NA,ALM_Air_Gate_Failed_Open_Bin15,Bin_Transfer_Pause,Clean_Batch_Status,Treat_Batch_Status,Transfer_Batch_Status,_700G_OPEN,_700G_CLOSE,Belt[4].Running,Manual_Mode,RemoteAndcoAnalogIn[15]);
   18: Loadout_Bin_Control(Bin_Loadout_Control[16],Loadout_Bin[16],O9_000_Bit00,Bin_Treat_Pause,Bin_Clean_Pause,TMR_Max_Treat_Delay,TMR_Max_Clean_Delay,I1_000_Bit00,NA,0,1,I4_000_Bit11,ALM_Air_Gate_Failed_Open_Bin16,Bin_Transfer_Pause,Clean_Batch_Status,Treat_Batch_Status,Transfer_Batch_Status,O9_000_Bit02,O9_000_Bit01,Belt[10].Running,Manual_Mode,R2S0_AENTR:3:I.Channel_0_Data);
